DATA_BLOCK "HMI"   // DB2
{ S7_Optimized_Access := 'TRUE' }
VERSION : 0.1
   VAR
      barcode : "Barcode Screen";
      networkHealth : "Network Health Screen";
      partCall : "Part Call Screen";
      screenNumber : Int;
      settings : "Settings";
      simStations : "Simulated Stations";
      tableNav : "Table Nav: HMI";
   END_VAR
BEGIN
END_DATA_BLOCK

DATA_BLOCK "PN Text Library"   // DB3
{ S7_Optimized_Access := 'TRUE' }
VERSION : 0.1
BEGIN
   pnText[0] := WSTRING#'';
   pnText[1] := WSTRING#'11.52.001.0545.000B';
   pnText[2] := WSTRING#'11.52.001.315.000B';
   pnText[3] := WSTRING#'11.52.001.316.001D';
   pnText[4] := WSTRING#'11.54.007.045.015D';
   pnText[5] := WSTRING#'11.54.007.052.007B';
   pnText[6] := WSTRING#'11.54.007.052.008A';
   pnText[7] := WSTRING#'11.54.007.052.009B';
   pnText[8] := WSTRING#'11.54.007.052.010B';
   pnText[9] := WSTRING#'11.54.007.315.026G';
   pnText[10] := WSTRING#'11.54.017.315.001F';
   pnText[11] := WSTRING#'16.08.208.011.010G';
   pnText[12] := WSTRING#'16.08.208.021.020C';
   pnText[13] := WSTRING#'16.08.208.031.020C';
   pnText[14] := WSTRING#'16.08.208.041.000A';
   pnText[15] := WSTRING#'16.08.208.051.000A';
   pnText[16] := WSTRING#'16.08.208.081.010B';
   pnText[17] := WSTRING#'16.08.208.091.000A';
   pnText[18] := WSTRING#'16.08.208.101.010C';
   pnText[19] := WSTRING#'16.08.208.111.000B';
   pnText[20] := WSTRING#'16.08.208.131.010L';
   pnText[21] := WSTRING#'16.08.208.151.010F';
   pnText[22] := WSTRING#'16.08.208.161.020F';
   pnText[23] := WSTRING#'16.08.208.301.000F';
   pnText[24] := WSTRING#'16.08.208.311.000F';
   pnText[25] := WSTRING#'16.08.208.321.000G';
   pnText[26] := WSTRING#'16.08.208.331.000F';
   pnText[27] := WSTRING#'16.08.208.411.030C';
   pnText[28] := WSTRING#'16.08.208.501.000B';
   pnText[29] := WSTRING#'16.08.208.531.020L';
   pnText[30] := WSTRING#'16.08.208.621.010C';
   pnText[31] := WSTRING#'16.08.208.631.000F';
   pnText[32] := WSTRING#'16.08.208.651.010B';
   pnText[33] := WSTRING#'16.08.208.661.000F';
   pnText[34] := WSTRING#'16.08.208.691.010D';
   pnText[35] := WSTRING#'16.08.209.031.010C';
   pnText[36] := WSTRING#'16.08.209.031.030B';
   pnText[37] := WSTRING#'16.08.209.031.050A';
   pnText[38] := WSTRING#'16.08.209.091.010C';
   pnText[39] := WSTRING#'16.08.209.091.030D';
   pnText[40] := WSTRING#'16.08.209.091.060A';
   pnText[41] := WSTRING#'16.08.209.232.010C';
   pnText[42] := WSTRING#'16.08.210.031.010B';
   pnText[43] := WSTRING#'16.08.210.421.010A';
   pnText[44] := WSTRING#'16.08.210.421.020A';
   pnText[45] := WSTRING#'16.08.210.421.030A';
   pnText[46] := WSTRING#'16.08.211.121.000G';
   pnText[47] := WSTRING#'16.08.211.291.000A';
   pnText[48] := WSTRING#'16.08.211.511.020F';
   pnText[49] := WSTRING#'16.08.211.551.000B';
   pnText[50] := WSTRING#'16.08.211.781.000A';
   pnText[51] := WSTRING#'16.08.211.801.010A';
   pnText[52] := WSTRING#'16.08.211.801.020A';
   pnText[53] := WSTRING#'16.08.211.806.020A';
   pnText[54] := WSTRING#'16.08.215.141.010C';
   pnText[55] := WSTRING#'16.08.215.871.010C';
   pnText[56] := WSTRING#'16.08.216.011.030B';
   pnText[57] := WSTRING#'16.08.216.053.000A';
   pnText[58] := WSTRING#'16.08.216.057.001A';
   pnText[59] := WSTRING#'16.08.216.141.010C';
   pnText[60] := WSTRING#'16.08.216.151.010B';
   pnText[61] := WSTRING#'16.08.216.161.020A';
   pnText[62] := WSTRING#'16.08.216.181.010B';
   pnText[63] := WSTRING#'16.08.216.181.090A';
   pnText[64] := WSTRING#'16.08.216.181.100A';
   pnText[65] := WSTRING#'16.08.216.181.110B';
   pnText[66] := WSTRING#'16.08.216.200.050A';
   pnText[67] := WSTRING#'16.08.216.202.080A';
   pnText[68] := WSTRING#'16.08.216.231.000B';
   pnText[69] := WSTRING#'16.08.216.251.000B';
   pnText[70] := WSTRING#'16.08.216.291.000A';
   pnText[71] := WSTRING#'16.08.216.315.000A';
   pnText[72] := WSTRING#'16.08.216.315.001A';
   pnText[73] := WSTRING#'16.08.216.315.002A';
   pnText[74] := WSTRING#'16.08.216.501.000C';
   pnText[75] := WSTRING#'16.08.216.501.010A';
   pnText[76] := WSTRING#'16.08.216.511.000C';
   pnText[77] := WSTRING#'16.08.216.515.008C';
   pnText[78] := WSTRING#'16.08.216.521.000C';
   pnText[79] := WSTRING#'16.08.216.526.002C';
   pnText[80] := WSTRING#'16.08.216.526.009A';
   pnText[81] := WSTRING#'16.08.216.551.000B';
   pnText[82] := WSTRING#'16.08.216.722.001A';
   pnText[83] := WSTRING#'16.08.216.790.001A';
   pnText[84] := WSTRING#'16.08.216.806.020A';
   pnText[85] := WSTRING#'16.08.216.831.020A';
   pnText[86] := WSTRING#'16.08.216.871.010C';
   pnText[87] := WSTRING#'16.08.216.910.020B';
   pnText[88] := WSTRING#'16.08.216.911.000C';
   pnText[89] := WSTRING#'16.08.216.911.000G';
   pnText[90] := WSTRING#'16.08.216.911.000H';
   pnText[91] := WSTRING#'16.08.216.911.030B';
   pnText[92] := WSTRING#'16.08.216.911.040B';
   pnText[93] := WSTRING#'16.08.216.912.050A';
   pnText[94] := WSTRING#'16.08.216.912.060B';
   pnText[95] := WSTRING#'16.08.216.951.010A';
   pnText[96] := WSTRING#'16.08.216.181.020A';
   pnText[97] := WSTRING#'16.08.217.411.080A';
   pnText[98] := WSTRING#'16.08.217.421.010A';
   pnText[99] := WSTRING#'16.08.217.421.130A';
   pnText[100] := WSTRING#'16.18.007.301.010A';
   pnText[101] := WSTRING#'16.18.007.301.020A';
   pnText[102] := WSTRING#'16.18.007.311.010A';
   pnText[103] := WSTRING#'16.18.007.311.020A';
   pnText[104] := WSTRING#'16.18.007.321.010B';
   pnText[105] := WSTRING#'16.18.008.301.010A';
   pnText[106] := WSTRING#'16.18.008.301.020A';
   pnText[107] := WSTRING#'16.18.008.301.030A';
   pnText[108] := WSTRING#'16.18.008.311.010A';
   pnText[109] := WSTRING#'16.18.008.311.020B';
   pnText[110] := WSTRING#'16.18.009.301.010A';
   pnText[111] := WSTRING#'16.18.009.301.020B';
   pnText[112] := WSTRING#'16.18.009.301.030A';
   pnText[113] := WSTRING#'16.18.009.301.040B';
   pnText[114] := WSTRING#'16.18.009.301.050A';
   pnText[115] := WSTRING#'16.18.009.311.010A';
   pnText[116] := WSTRING#'16.18.009.321.010A';
   pnText[117] := WSTRING#'16.18.009.321.020B';
   pnText[118] := WSTRING#'16.18.009.321.030A';
   pnText[119] := WSTRING#'16.18.009.331.030A';
   pnText[120] := WSTRING#'16.18.009.331.050A';
   pnText[121] := WSTRING#'16.18.009.371.010A';
   pnText[122] := WSTRING#'16.18.011.301.010A';
   pnText[123] := WSTRING#'16.18.011.301.020B';
   pnText[124] := WSTRING#'16.18.011.301.030A';
   pnText[125] := WSTRING#'16.18.011.301.040B';
   pnText[126] := WSTRING#'16.18.011.311.020A';
   pnText[127] := WSTRING#'16.18.011.321.010A';
   pnText[128] := WSTRING#'16.18.011.321.020B';
   pnText[129] := WSTRING#'16.18.011.321.030A';
   pnText[130] := WSTRING#'16.18.011.331.010A';
   pnText[131] := WSTRING#'16.18.011.331.020D';
   pnText[132] := WSTRING#'16.18.012.401.010A';
   pnText[133] := WSTRING#'16.18.012.401.020A';
   pnText[134] := WSTRING#'16.18.012.411.010A';
   pnText[135] := WSTRING#'16.18.012.411.020B';
   pnText[136] := WSTRING#'16.18.012.431.010A';
   pnText[137] := WSTRING#'16.18.012.441.010A';
   pnText[138] := WSTRING#'16.18.013.411.010A';
   pnText[139] := WSTRING#'16.18.013.411.020B';
   pnText[140] := WSTRING#'16.18.013.411.030A';
   pnText[141] := WSTRING#'16.18.013.421.010A';
   pnText[142] := WSTRING#'16.18.014.411.010A';
   pnText[143] := WSTRING#'16.18.014.411.030A';
   pnText[144] := WSTRING#'16.18.015.401.010A';
   pnText[145] := WSTRING#'16.18.015.411.010A';
   pnText[146] := WSTRING#'16.18.015.411.020B';
   pnText[147] := WSTRING#'16.18.015.411.030A';
   pnText[148] := WSTRING#'16.18.015.421.010A';
   pnText[149] := WSTRING#'16.18.015.421.020B';
   pnText[150] := WSTRING#'16.18.017.301.010A';
   pnText[151] := WSTRING#'16.18.017.301.020A';
   pnText[152] := WSTRING#'16.18.017.301.030A';
   pnText[153] := WSTRING#'16.18.017.301.040A';
   pnText[154] := WSTRING#'16.18.017.301.050A';
   pnText[155] := WSTRING#'16.18.017.311.010A';
   pnText[156] := WSTRING#'16.18.017.321.010A';
   pnText[157] := WSTRING#'16.18.017.321.020A';
   pnText[158] := WSTRING#'16.18.018.400.000A';
   pnText[159] := WSTRING#'16.18.018.401.010A';
   pnText[160] := WSTRING#'16.18.018.401.020B';
   pnText[161] := WSTRING#'16.18.018.401.030A';
   pnText[162] := WSTRING#'16.18.018.411.010A';
   pnText[163] := WSTRING#'16.18.018.421.010B';
   pnText[164] := WSTRING#'16.32.112.054.041A';
   pnText[165] := WSTRING#'16.32.112.057.010A';
   pnText[166] := WSTRING#'16.32.112.500.060D';
   pnText[167] := WSTRING#'16.32.112.500.090B';
   pnText[168] := WSTRING#'16.32.112.500.100A';
   pnText[169] := WSTRING#'16.32.112.500.120A';
   pnText[170] := WSTRING#'16.32.112.500.150B';
   pnText[171] := WSTRING#'16.32.112.500.160A';
   pnText[172] := WSTRING#'16.32.112.500.220A';
   pnText[173] := WSTRING#'16.32.112.500.300E';
   pnText[174] := WSTRING#'16.32.112.500.520B';
   pnText[175] := WSTRING#'16.32.112.502.050B';
   pnText[176] := WSTRING#'16.32.112.502.060B';
   pnText[177] := WSTRING#'16.32.112.502.070E';
   pnText[178] := WSTRING#'16.32.112.503.210A';
   pnText[179] := WSTRING#'16.32.112.503.220A';
   pnText[180] := WSTRING#'16.32.112.504.060A';
   pnText[181] := WSTRING#'16.32.112.504.070G';
   pnText[182] := WSTRING#'16.32.112.509.050E';
   pnText[183] := WSTRING#'16.32.112.509.070A';
   pnText[184] := WSTRING#'16.32.112.509.080F';
   pnText[185] := WSTRING#'16.32.112.516.110E';
   pnText[186] := WSTRING#'16.32.112.520.300E';
   pnText[187] := WSTRING#'16.32.112.521.010B';
   pnText[188] := WSTRING#'16.32.112.521.020B';
   pnText[189] := WSTRING#'16.32.112.521.030A';
   pnText[190] := WSTRING#'16.32.112.522.040D';
   pnText[191] := WSTRING#'16.32.112.522.050A';
   pnText[192] := WSTRING#'16.32.112.522.130A';
   pnText[193] := WSTRING#'16.32.112.529.010A';
   pnText[194] := WSTRING#'16.32.112.529.020B';
   pnText[195] := WSTRING#'16.32.112.529.030A';
   pnText[196] := WSTRING#'16.32.112.529.050D';
   pnText[197] := WSTRING#'16.32.112.536.010A';
   pnText[198] := WSTRING#'16.32.112.543.020A';
   pnText[199] := WSTRING#'16.32.112.543.210E';
   pnText[200] := WSTRING#'16.32.112.553.010A';
   pnText[201] := WSTRING#'16.32.112.553.020A';
   pnText[202] := WSTRING#'16.32.112.553.100D';
   pnText[203] := WSTRING#'16.32.112.553.220A';
   pnText[204] := WSTRING#'16.32.112.580.020A';
   pnText[205] := WSTRING#'16.32.112.601.030A';
   pnText[206] := WSTRING#'16.32.112.601.040A';
   pnText[207] := WSTRING#'16.32.112.621.010A';
   pnText[208] := WSTRING#'16.32.112.621.020A';
   pnText[209] := WSTRING#'16.32.112.704.000C';
   pnText[210] := WSTRING#'16.32.112.751.000D';
   pnText[211] := WSTRING#'16.32.112.751.001C';
   pnText[212] := WSTRING#'16.32.112.757.000A';
   pnText[213] := WSTRING#'16.32.112.757.001A';
   pnText[214] := WSTRING#'16.32.112.851.000A';
   pnText[215] := WSTRING#'16.32.112.851.001A';
   pnText[216] := WSTRING#'16.32.112.870.000C';
   pnText[217] := WSTRING#'16.32.307.211.150B';
   pnText[218] := WSTRING#'16.32.307.211.170B';
   pnText[219] := WSTRING#'16.32.307.212.320C';
   pnText[220] := WSTRING#'16.32.307.232.300B';
   pnText[221] := WSTRING#'16.32.307.262.300B';
   pnText[222] := WSTRING#'16.32.307.312.310A';
   pnText[223] := WSTRING#'16.32.307.461.160A';
   pnText[224] := WSTRING#'16.32.407.241.150B';
   pnText[225] := WSTRING#'16.32.407.241.170B';
   pnText[226] := WSTRING#'16.32.407.441.160A';
   pnText[227] := WSTRING#'16.32.606.311.010C';
   pnText[228] := WSTRING#'16.32.606.311.040B';
   pnText[229] := WSTRING#'16.32.606.311.050B';
   pnText[230] := WSTRING#'16.32.606.311.060A';
   pnText[231] := WSTRING#'16.32.606.311.070A';
   pnText[232] := WSTRING#'16.32.606.321.010B';
   pnText[233] := WSTRING#'16.32.606.321.030B';
   pnText[234] := WSTRING#'16.32.706.311.010C';
   pnText[235] := WSTRING#'16.32.706.311.020B';
   pnText[236] := WSTRING#'16.32.706.311.040B';
   pnText[237] := WSTRING#'16.32.706.311.050B';
   pnText[238] := WSTRING#'16.32.706.321.010B';
   pnText[239] := WSTRING#'16.32.706.321.030B';
   pnText[240] := WSTRING#'16.32.706.401.040A';
   pnText[241] := WSTRING#'16.32.706.401.050A';
   pnText[242] := WSTRING#'16.32.806.502.080A';
   pnText[243] := WSTRING#'DUNNAGE';
   pnText[244] := WSTRING#'PEANUTS';
   pnText[245] := WSTRING#'RINGS CART';
END_DATA_BLOCK

DATA_BLOCK "LED Sign"   // DB4
{ S7_Optimized_Access := 'TRUE' }
VERSION : 0.1
   VAR
      request : "LED Sign Data";
   END_VAR
BEGIN
END_DATA_BLOCK

DATA_BLOCK "Recipe Buffer"   // DB5
{ S7_Optimized_Access := 'TRUE' }
VERSION : 0.1
BEGIN
END_DATA_BLOCK

DATA_BLOCK "HMI Stations"   // DB6
{ S7_Optimized_Access := 'TRUE' }
VERSION : 0.1
   VAR
      me : Array[0.."hmiStnCount"] of "HMIS: Compressed";
   END_VAR
BEGIN
END_DATA_BLOCK

DATA_BLOCK "Stations"   // DB10
{ S7_Optimized_Access := 'TRUE' }
VERSION : 0.1
BEGIN
   stn[0].id.dropZone := 1;
   stn[0].id.lineName := WSTRING#'VOLVO 16';
   stn[0].ioData.kp8.output := 16#0000_0000;
   stn[0].ioData.stkLight := 16#0000_0000;
   stn[0].wipData."name" := WSTRING#'';
   stn[1].id.dropZone := 2;
   stn[1].id.lineName := WSTRING#'VOLVO 16';
   stn[1].ioData.kp8.output := 16#0000_0000;
   stn[1].ioData.stkLight := 16#0000_0000;
   stn[1].wipData."name" := WSTRING#'';
   stn[2].id.dropZone := 3;
   stn[2].id.lineName := WSTRING#'VOLVO 16';
   stn[2].ioData.kp8.output := 16#0000_0000;
   stn[2].ioData.stkLight := 16#0000_0000;
   stn[2].wipData."name" := WSTRING#'';
   stn[3].id.dropZone := 4;
   stn[3].id.lineName := WSTRING#'VOLVO 16';
   stn[3].ioData.kp8.output := 16#0000_0000;
   stn[3].ioData.stkLight := 16#0000_0000;
   stn[3].wipData."name" := WSTRING#'';
   stn[4].id.lineName := WSTRING#'';
   stn[4].ioData.kp8.output := 16#0000_0000;
   stn[4].ioData.stkLight := 16#0000_0000;
   stn[4].wipData."name" := WSTRING#'';
   stn[5].id.lineName := WSTRING#'';
   stn[5].ioData.kp8.output := 16#0000_0000;
   stn[5].ioData.stkLight := 16#0000_0000;
   stn[5].wipData."name" := WSTRING#'';
   stn[6].id.lineName := WSTRING#'';
   stn[6].ioData.kp8.output := 16#0000_0000;
   stn[6].ioData.stkLight := 16#0000_0000;
   stn[6].wipData."name" := WSTRING#'';
   stn[7].id.lineName := WSTRING#'';
   stn[7].ioData.kp8.output := 16#0000_0000;
   stn[7].ioData.stkLight := 16#0000_0000;
   stn[7].wipData."name" := WSTRING#'';
   stn[8].id.lineName := WSTRING#'';
   stn[8].ioData.kp8.output := 16#0000_0000;
   stn[8].ioData.stkLight := 16#0000_0000;
   stn[8].wipData."name" := WSTRING#'';
   stn[9].id.lineName := WSTRING#'';
   stn[9].ioData.kp8.output := 16#0000_0000;
   stn[9].ioData.stkLight := 16#0000_0000;
   stn[9].wipData."name" := WSTRING#'';
   stn[10].id.lineName := WSTRING#'';
   stn[10].ioData.kp8.output := 16#0000_0000;
   stn[10].ioData.stkLight := 16#0000_0000;
   stn[10].wipData."name" := WSTRING#'';
   stn[11].id.lineName := WSTRING#'';
   stn[11].ioData.kp8.output := 16#0000_0000;
   stn[11].ioData.stkLight := 16#0000_0000;
   stn[11].wipData."name" := WSTRING#'';
   stn[12].id.lineName := WSTRING#'';
   stn[12].ioData.kp8.output := 16#0000_0000;
   stn[12].ioData.stkLight := 16#0000_0000;
   stn[12].wipData."name" := WSTRING#'';
   stn[13].id.lineName := WSTRING#'';
   stn[13].ioData.kp8.output := 16#0000_0000;
   stn[13].ioData.stkLight := 16#0000_0000;
   stn[13].wipData."name" := WSTRING#'';
   stn[14].id.lineName := WSTRING#'';
   stn[14].ioData.kp8.output := 16#0000_0000;
   stn[14].ioData.stkLight := 16#0000_0000;
   stn[14].wipData."name" := WSTRING#'';
   stn[15].id.lineName := WSTRING#'';
   stn[15].ioData.kp8.output := 16#0000_0000;
   stn[15].ioData.stkLight := 16#0000_0000;
   stn[15].wipData."name" := WSTRING#'';
   stn[16].id.lineName := WSTRING#'';
   stn[16].ioData.kp8.output := 16#0000_0000;
   stn[16].ioData.stkLight := 16#0000_0000;
   stn[16].wipData."name" := WSTRING#'';
   stn[17].id.lineName := WSTRING#'';
   stn[17].ioData.kp8.output := 16#0000_0000;
   stn[17].ioData.stkLight := 16#0000_0000;
   stn[17].wipData."name" := WSTRING#'';
   stn[18].id.lineName := WSTRING#'';
   stn[18].ioData.kp8.output := 16#0000_0000;
   stn[18].ioData.stkLight := 16#0000_0000;
   stn[18].wipData."name" := WSTRING#'';
   stn[19].id.lineName := WSTRING#'';
   stn[19].ioData.kp8.output := 16#0000_0000;
   stn[19].ioData.stkLight := 16#0000_0000;
   stn[19].wipData."name" := WSTRING#'';
   stn[20].id.lineName := WSTRING#'';
   stn[20].ioData.kp8.output := 16#0000_0000;
   stn[20].ioData.stkLight := 16#0000_0000;
   stn[20].wipData."name" := WSTRING#'';
   stn[21].id.lineName := WSTRING#'';
   stn[21].ioData.kp8.output := 16#0000_0000;
   stn[21].ioData.stkLight := 16#0000_0000;
   stn[21].wipData."name" := WSTRING#'';
   stn[22].id.lineName := WSTRING#'';
   stn[22].ioData.kp8.output := 16#0000_0000;
   stn[22].ioData.stkLight := 16#0000_0000;
   stn[22].wipData."name" := WSTRING#'';
   stn[23].id.lineName := WSTRING#'';
   stn[23].ioData.kp8.output := 16#0000_0000;
   stn[23].ioData.stkLight := 16#0000_0000;
   stn[23].wipData."name" := WSTRING#'';
   stn[24].id.lineName := WSTRING#'';
   stn[24].ioData.kp8.output := 16#0000_0000;
   stn[24].ioData.stkLight := 16#0000_0000;
   stn[24].wipData."name" := WSTRING#'';
   stn[25].id.lineName := WSTRING#'';
   stn[25].ioData.kp8.output := 16#0000_0000;
   stn[25].ioData.stkLight := 16#0000_0000;
   stn[25].wipData."name" := WSTRING#'';
   stn[26].id.lineName := WSTRING#'';
   stn[26].ioData.kp8.output := 16#0000_0000;
   stn[26].ioData.stkLight := 16#0000_0000;
   stn[26].wipData."name" := WSTRING#'';
   stn[27].id.lineName := WSTRING#'';
   stn[27].ioData.kp8.output := 16#0000_0000;
   stn[27].ioData.stkLight := 16#0000_0000;
   stn[27].wipData."name" := WSTRING#'';
   stn[28].id.lineName := WSTRING#'';
   stn[28].ioData.kp8.output := 16#0000_0000;
   stn[28].ioData.stkLight := 16#0000_0000;
   stn[28].wipData."name" := WSTRING#'';
   stn[29].id.lineName := WSTRING#'';
   stn[29].ioData.kp8.output := 16#0000_0000;
   stn[29].ioData.stkLight := 16#0000_0000;
   stn[29].wipData."name" := WSTRING#'';
   stn[30].id.lineName := WSTRING#'';
   stn[30].ioData.kp8.output := 16#0000_0000;
   stn[30].ioData.stkLight := 16#0000_0000;
   stn[30].wipData."name" := WSTRING#'';
   stn[31].id.lineName := WSTRING#'';
   stn[31].ioData.kp8.output := 16#0000_0000;
   stn[31].ioData.stkLight := 16#0000_0000;
   stn[31].wipData."name" := WSTRING#'';
   stn[32].id.lineName := WSTRING#'';
   stn[32].ioData.kp8.output := 16#0000_0000;
   stn[32].ioData.stkLight := 16#0000_0000;
   stn[32].wipData."name" := WSTRING#'';
   stn[33].id.lineName := WSTRING#'';
   stn[33].ioData.kp8.output := 16#0000_0000;
   stn[33].ioData.stkLight := 16#0000_0000;
   stn[33].wipData."name" := WSTRING#'';
   stn[34].id.lineName := WSTRING#'';
   stn[34].ioData.kp8.output := 16#0000_0000;
   stn[34].ioData.stkLight := 16#0000_0000;
   stn[34].wipData."name" := WSTRING#'';
   stn[35].id.lineName := WSTRING#'';
   stn[35].ioData.kp8.output := 16#0000_0000;
   stn[35].ioData.stkLight := 16#0000_0000;
   stn[35].wipData."name" := WSTRING#'';
   stn[36].id.lineName := WSTRING#'';
   stn[36].ioData.kp8.output := 16#0000_0000;
   stn[36].ioData.stkLight := 16#0000_0000;
   stn[36].wipData."name" := WSTRING#'';
   stn[37].id.lineName := WSTRING#'';
   stn[37].ioData.kp8.output := 16#0000_0000;
   stn[37].ioData.stkLight := 16#0000_0000;
   stn[37].wipData."name" := WSTRING#'';
   stn[38].id.lineName := WSTRING#'';
   stn[38].ioData.kp8.output := 16#0000_0000;
   stn[38].ioData.stkLight := 16#0000_0000;
   stn[38].wipData."name" := WSTRING#'';
END_DATA_BLOCK

DATA_BLOCK "Part Requests"   // DB11
{ S7_Optimized_Access := 'TRUE' }
VERSION : 0.1
BEGIN
END_DATA_BLOCK

DATA_BLOCK "PN Code Library"   // DB12
{ S7_Optimized_Access := 'TRUE' }
VERSION : 0.1
BEGIN
   stn[0].wipBtn[0,0] := 0;
   stn[0].wipBtn[0,1] := 0;
   stn[0].wipBtn[0,2] := 0;
   stn[0].wipBtn[0,4] := 0;
   stn[0].wipBtn[0,5] := 0;
   stn[0].wipBtn[0,6] := 0;
   stn[0].wipBtn[1,0] := 0;
   stn[0].wipBtn[1,1] := 0;
   stn[0].wipBtn[1,2] := 0;
   stn[0].wipBtn[1,3] := 0;
   stn[0].wipBtn[1,4] := 0;
   stn[0].wipBtn[1,5] := 0;
   stn[0].wipBtn[1,6] := 0;
   stn[0].wipBtn[1,7] := 0;
   stn[0].wipBtn[2,0] := 0;
   stn[0].wipBtn[2,1] := 0;
   stn[0].wipBtn[2,2] := 0;
   stn[0].wipBtn[2,3] := 0;
   stn[0].wipBtn[2,4] := 0;
   stn[0].wipBtn[2,5] := 0;
   stn[0].wipBtn[2,6] := 0;
   stn[0].wipBtn[2,7] := 0;
   stn[0].wipBtn[3,0] := 0;
   stn[0].wipBtn[3,1] := 0;
   stn[0].wipBtn[3,2] := 0;
   stn[0].wipBtn[3,3] := 0;
   stn[0].wipBtn[3,4] := 0;
   stn[0].wipBtn[3,5] := 0;
   stn[0].wipBtn[3,6] := 0;
   stn[0].wipBtn[3,7] := 0;
   stn[0].wipBtn[4,0] := 0;
   stn[0].wipBtn[4,1] := 0;
   stn[0].wipBtn[4,2] := 0;
   stn[0].wipBtn[4,3] := 0;
   stn[0].wipBtn[4,4] := 0;
   stn[0].wipBtn[4,5] := 0;
   stn[0].wipBtn[4,6] := 0;
   stn[0].wipBtn[4,7] := 0;
   stn[0].wipBtn[5,0] := 0;
   stn[0].wipBtn[5,1] := 0;
   stn[0].wipBtn[5,2] := 0;
   stn[0].wipBtn[5,3] := 0;
   stn[0].wipBtn[5,4] := 0;
   stn[0].wipBtn[5,5] := 0;
   stn[0].wipBtn[5,6] := 0;
   stn[0].wipBtn[5,7] := 0;
   stn[0].wipBtn[6,0] := 0;
   stn[0].wipBtn[6,1] := 0;
   stn[0].wipBtn[6,2] := 0;
   stn[0].wipBtn[6,3] := 0;
   stn[0].wipBtn[6,4] := 0;
   stn[0].wipBtn[6,5] := 0;
   stn[0].wipBtn[6,6] := 0;
   stn[0].wipBtn[6,7] := 0;
   stn[0].wipBtn[7,0] := 0;
   stn[0].wipBtn[7,1] := 0;
   stn[0].wipBtn[7,2] := 0;
   stn[0].wipBtn[7,3] := 0;
   stn[0].wipBtn[7,4] := 0;
   stn[0].wipBtn[7,5] := 0;
   stn[0].wipBtn[7,6] := 0;
   stn[0].wipBtn[7,7] := 0;
   stn[0].wipBtn[8,0] := 0;
   stn[0].wipBtn[8,1] := 0;
   stn[0].wipBtn[8,2] := 0;
   stn[0].wipBtn[8,3] := 0;
   stn[0].wipBtn[8,4] := 0;
   stn[0].wipBtn[8,5] := 0;
   stn[0].wipBtn[8,6] := 0;
   stn[0].wipBtn[8,7] := 0;
   stn[0].wipBtn[9,0] := 0;
   stn[0].wipBtn[9,1] := 0;
   stn[0].wipBtn[9,2] := 0;
   stn[0].wipBtn[9,3] := 0;
   stn[0].wipBtn[9,4] := 0;
   stn[0].wipBtn[9,5] := 0;
   stn[0].wipBtn[9,6] := 0;
   stn[0].wipBtn[9,7] := 0;
   stn[0].wipBtn[10,0] := 0;
   stn[0].wipBtn[10,1] := 0;
   stn[0].wipBtn[10,2] := 0;
   stn[0].wipBtn[10,3] := 0;
   stn[0].wipBtn[10,4] := 0;
   stn[0].wipBtn[10,5] := 0;
   stn[0].wipBtn[10,6] := 0;
   stn[0].wipBtn[10,7] := 0;
   stn[0].wipBtn[11,0] := 0;
   stn[0].wipBtn[11,1] := 0;
   stn[0].wipBtn[11,2] := 0;
   stn[0].wipBtn[11,3] := 0;
   stn[0].wipBtn[11,4] := 0;
   stn[0].wipBtn[11,5] := 0;
   stn[0].wipBtn[11,6] := 0;
   stn[0].wipBtn[11,7] := 0;
   stn[0].wipBtn[12,0] := 0;
   stn[0].wipBtn[12,1] := 0;
   stn[0].wipBtn[12,2] := 0;
   stn[0].wipBtn[12,3] := 0;
   stn[0].wipBtn[12,4] := 0;
   stn[0].wipBtn[12,5] := 0;
   stn[0].wipBtn[12,6] := 0;
   stn[0].wipBtn[12,7] := 0;
   stn[0].wipBtn[13,0] := 0;
   stn[0].wipBtn[13,1] := 0;
   stn[0].wipBtn[13,2] := 0;
   stn[0].wipBtn[13,3] := 0;
   stn[0].wipBtn[13,4] := 0;
   stn[0].wipBtn[13,5] := 0;
   stn[0].wipBtn[13,6] := 0;
   stn[0].wipBtn[13,7] := 0;
   stn[0].wipBtn[14,0] := 0;
   stn[0].wipBtn[14,1] := 0;
   stn[0].wipBtn[14,2] := 0;
   stn[0].wipBtn[14,3] := 0;
   stn[0].wipBtn[14,4] := 0;
   stn[0].wipBtn[14,5] := 0;
   stn[0].wipBtn[14,6] := 0;
   stn[0].wipBtn[14,7] := 0;
   stn[0].wipBtn[15,0] := 0;
   stn[0].wipBtn[15,1] := 0;
   stn[0].wipBtn[15,2] := 0;
   stn[0].wipBtn[15,3] := 0;
   stn[0].wipBtn[15,4] := 0;
   stn[0].wipBtn[15,5] := 0;
   stn[0].wipBtn[15,6] := 0;
   stn[0].wipBtn[15,7] := 0;
   stn[0].wipBtn[16,0] := 0;
   stn[0].wipBtn[16,1] := 0;
   stn[0].wipBtn[16,2] := 0;
   stn[0].wipBtn[16,3] := 0;
   stn[0].wipBtn[16,4] := 0;
   stn[0].wipBtn[16,5] := 0;
   stn[0].wipBtn[16,6] := 0;
   stn[0].wipBtn[16,7] := 0;
   stn[0].wipBtn[17,0] := 0;
   stn[0].wipBtn[17,1] := 0;
   stn[0].wipBtn[17,2] := 0;
   stn[0].wipBtn[17,3] := 0;
   stn[0].wipBtn[17,4] := 0;
   stn[0].wipBtn[17,5] := 0;
   stn[0].wipBtn[17,6] := 0;
   stn[0].wipBtn[17,7] := 0;
   stn[0].wipBtn[18,0] := 0;
   stn[0].wipBtn[18,1] := 0;
   stn[0].wipBtn[18,2] := 0;
   stn[0].wipBtn[18,3] := 0;
   stn[0].wipBtn[18,4] := 0;
   stn[0].wipBtn[18,5] := 0;
   stn[0].wipBtn[18,6] := 0;
   stn[0].wipBtn[18,7] := 0;
   stn[0].wipBtn[19,0] := 0;
   stn[0].wipBtn[19,1] := 0;
   stn[0].wipBtn[19,2] := 0;
   stn[0].wipBtn[19,3] := 0;
   stn[0].wipBtn[19,4] := 0;
   stn[0].wipBtn[19,5] := 0;
   stn[0].wipBtn[19,6] := 0;
   stn[0].wipBtn[19,7] := 0;
   stn[0].wipBtn[20,0] := 0;
   stn[0].wipBtn[20,1] := 0;
   stn[0].wipBtn[20,2] := 0;
   stn[0].wipBtn[20,3] := 0;
   stn[0].wipBtn[20,4] := 0;
   stn[0].wipBtn[20,5] := 0;
   stn[0].wipBtn[20,6] := 0;
   stn[0].wipBtn[20,7] := 0;
   stn[0].wipBtn[21,0] := 0;
   stn[0].wipBtn[21,1] := 0;
   stn[0].wipBtn[21,2] := 0;
   stn[0].wipBtn[21,3] := 0;
   stn[0].wipBtn[21,4] := 0;
   stn[0].wipBtn[21,5] := 0;
   stn[0].wipBtn[21,6] := 0;
   stn[0].wipBtn[21,7] := 0;
   stn[0].wipBtn[22,0] := 0;
   stn[0].wipBtn[22,1] := 0;
   stn[0].wipBtn[22,2] := 0;
   stn[0].wipBtn[22,3] := 0;
   stn[0].wipBtn[22,4] := 0;
   stn[0].wipBtn[22,5] := 0;
   stn[0].wipBtn[22,6] := 0;
   stn[0].wipBtn[22,7] := 0;
   stn[0].wipBtn[23,0] := 0;
   stn[0].wipBtn[23,1] := 0;
   stn[0].wipBtn[23,2] := 0;
   stn[0].wipBtn[23,3] := 0;
   stn[0].wipBtn[23,4] := 0;
   stn[0].wipBtn[23,5] := 0;
   stn[0].wipBtn[23,6] := 0;
   stn[0].wipBtn[23,7] := 0;
   stn[0].wipBtn[24,0] := 0;
   stn[0].wipBtn[24,1] := 0;
   stn[0].wipBtn[24,2] := 0;
   stn[0].wipBtn[24,3] := 0;
   stn[0].wipBtn[24,4] := 0;
   stn[0].wipBtn[24,5] := 0;
   stn[0].wipBtn[24,6] := 0;
   stn[0].wipBtn[24,7] := 0;
   stn[0].wipBtn[25,0] := 0;
   stn[0].wipBtn[25,1] := 0;
   stn[0].wipBtn[25,2] := 0;
   stn[0].wipBtn[25,3] := 0;
   stn[0].wipBtn[25,4] := 0;
   stn[0].wipBtn[25,5] := 0;
   stn[0].wipBtn[25,6] := 0;
   stn[0].wipBtn[25,7] := 0;
   stn[0].wipBtn[26,0] := 0;
   stn[0].wipBtn[26,1] := 0;
   stn[0].wipBtn[26,2] := 0;
   stn[0].wipBtn[26,3] := 0;
   stn[0].wipBtn[26,4] := 0;
   stn[0].wipBtn[26,5] := 0;
   stn[0].wipBtn[26,6] := 0;
   stn[0].wipBtn[26,7] := 0;
   stn[0].wipBtn[27,0] := 0;
   stn[0].wipBtn[27,1] := 0;
   stn[0].wipBtn[27,2] := 0;
   stn[0].wipBtn[27,3] := 0;
   stn[0].wipBtn[27,4] := 0;
   stn[0].wipBtn[27,5] := 0;
   stn[0].wipBtn[27,6] := 0;
   stn[0].wipBtn[27,7] := 0;
   stn[0].wipBtn[28,0] := 0;
   stn[0].wipBtn[28,1] := 0;
   stn[0].wipBtn[28,2] := 0;
   stn[0].wipBtn[28,3] := 0;
   stn[0].wipBtn[28,4] := 0;
   stn[0].wipBtn[28,5] := 0;
   stn[0].wipBtn[28,6] := 0;
   stn[0].wipBtn[28,7] := 0;
   stn[0].wipBtn[29,0] := 0;
   stn[0].wipBtn[29,1] := 0;
   stn[0].wipBtn[29,2] := 0;
   stn[0].wipBtn[29,3] := 0;
   stn[0].wipBtn[29,4] := 0;
   stn[0].wipBtn[29,5] := 0;
   stn[0].wipBtn[29,6] := 0;
   stn[0].wipBtn[29,7] := 0;
   stn[0].wipBtn[30,0] := 0;
   stn[0].wipBtn[30,1] := 0;
   stn[0].wipBtn[30,2] := 0;
   stn[0].wipBtn[30,3] := 0;
   stn[0].wipBtn[30,4] := 0;
   stn[0].wipBtn[30,5] := 0;
   stn[0].wipBtn[30,6] := 0;
   stn[0].wipBtn[30,7] := 0;
   stn[0].wipBtn[31,0] := 0;
   stn[0].wipBtn[31,1] := 0;
   stn[0].wipBtn[31,2] := 0;
   stn[0].wipBtn[31,3] := 0;
   stn[0].wipBtn[31,4] := 0;
   stn[0].wipBtn[31,5] := 0;
   stn[0].wipBtn[31,6] := 0;
   stn[0].wipBtn[31,7] := 0;
   stn[0].wipBtn[32,0] := 0;
   stn[0].wipBtn[32,1] := 0;
   stn[0].wipBtn[32,2] := 0;
   stn[0].wipBtn[32,3] := 0;
   stn[0].wipBtn[32,4] := 0;
   stn[0].wipBtn[32,5] := 0;
   stn[0].wipBtn[32,6] := 0;
   stn[0].wipBtn[32,7] := 0;
   stn[0].wipBtn[33,0] := 0;
   stn[0].wipBtn[33,1] := 0;
   stn[0].wipBtn[33,2] := 0;
   stn[0].wipBtn[33,3] := 0;
   stn[0].wipBtn[33,4] := 0;
   stn[0].wipBtn[33,5] := 0;
   stn[0].wipBtn[33,6] := 0;
   stn[0].wipBtn[33,7] := 0;
   stn[0].wipBtn[34,0] := 0;
   stn[0].wipBtn[34,1] := 0;
   stn[0].wipBtn[34,2] := 0;
   stn[0].wipBtn[34,3] := 0;
   stn[0].wipBtn[34,4] := 0;
   stn[0].wipBtn[34,5] := 0;
   stn[0].wipBtn[34,6] := 0;
   stn[0].wipBtn[34,7] := 0;
   stn[0].wipBtn[35,0] := 0;
   stn[0].wipBtn[35,1] := 0;
   stn[0].wipBtn[35,2] := 0;
   stn[0].wipBtn[35,3] := 0;
   stn[0].wipBtn[35,4] := 0;
   stn[0].wipBtn[35,5] := 0;
   stn[0].wipBtn[35,6] := 0;
   stn[0].wipBtn[35,7] := 0;
   stn[0].wipBtn[36,0] := 0;
   stn[0].wipBtn[36,1] := 0;
   stn[0].wipBtn[36,2] := 0;
   stn[0].wipBtn[36,3] := 0;
   stn[0].wipBtn[36,4] := 0;
   stn[0].wipBtn[36,5] := 0;
   stn[0].wipBtn[36,6] := 0;
   stn[0].wipBtn[36,7] := 0;
   stn[0].wipBtn[37,0] := 0;
   stn[0].wipBtn[37,1] := 0;
   stn[0].wipBtn[37,2] := 0;
   stn[0].wipBtn[37,3] := 0;
   stn[0].wipBtn[37,4] := 0;
   stn[0].wipBtn[37,5] := 0;
   stn[0].wipBtn[37,6] := 0;
   stn[0].wipBtn[37,7] := 0;
   stn[0].wipBtn[38,0] := 0;
   stn[0].wipBtn[38,1] := 0;
   stn[0].wipBtn[38,2] := 0;
   stn[0].wipBtn[38,3] := 0;
   stn[0].wipBtn[38,4] := 0;
   stn[0].wipBtn[38,5] := 0;
   stn[0].wipBtn[38,6] := 0;
   stn[0].wipBtn[38,7] := 0;
   stn[0].wipBtn[39,0] := 0;
   stn[0].wipBtn[39,1] := 0;
   stn[0].wipBtn[39,2] := 0;
   stn[0].wipBtn[39,3] := 0;
   stn[0].wipBtn[39,4] := 0;
   stn[0].wipBtn[39,5] := 0;
   stn[0].wipBtn[39,6] := 0;
   stn[0].wipBtn[39,7] := 0;
   stn[0].wipBtn[40,0] := 0;
   stn[0].wipBtn[40,1] := 0;
   stn[0].wipBtn[40,2] := 0;
   stn[0].wipBtn[40,3] := 0;
   stn[0].wipBtn[40,4] := 0;
   stn[0].wipBtn[40,5] := 0;
   stn[0].wipBtn[40,6] := 0;
   stn[0].wipBtn[40,7] := 0;
   stn[0].wipBtn[41,0] := 0;
   stn[0].wipBtn[41,1] := 0;
   stn[0].wipBtn[41,2] := 0;
   stn[0].wipBtn[41,3] := 0;
   stn[0].wipBtn[41,4] := 0;
   stn[0].wipBtn[41,5] := 0;
   stn[0].wipBtn[41,6] := 0;
   stn[0].wipBtn[41,7] := 0;
   stn[0].wipBtn[42,0] := 0;
   stn[0].wipBtn[42,1] := 0;
   stn[0].wipBtn[42,2] := 0;
   stn[0].wipBtn[42,3] := 0;
   stn[0].wipBtn[42,4] := 0;
   stn[0].wipBtn[42,5] := 0;
   stn[0].wipBtn[42,6] := 0;
   stn[0].wipBtn[42,7] := 0;
   stn[0].wipBtn[43,0] := 0;
   stn[0].wipBtn[43,1] := 0;
   stn[0].wipBtn[43,2] := 0;
   stn[0].wipBtn[43,3] := 0;
   stn[0].wipBtn[43,4] := 0;
   stn[0].wipBtn[43,5] := 0;
   stn[0].wipBtn[43,6] := 0;
   stn[0].wipBtn[43,7] := 0;
   stn[0].wipBtn[44,0] := 0;
   stn[0].wipBtn[44,1] := 0;
   stn[0].wipBtn[44,2] := 0;
   stn[0].wipBtn[44,3] := 0;
   stn[0].wipBtn[44,4] := 0;
   stn[0].wipBtn[44,5] := 0;
   stn[0].wipBtn[44,6] := 0;
   stn[0].wipBtn[44,7] := 0;
   stn[0].wipBtn[45,0] := 0;
   stn[0].wipBtn[45,1] := 0;
   stn[0].wipBtn[45,2] := 0;
   stn[0].wipBtn[45,3] := 0;
   stn[0].wipBtn[45,4] := 0;
   stn[0].wipBtn[45,5] := 0;
   stn[0].wipBtn[45,6] := 0;
   stn[0].wipBtn[45,7] := 0;
   stn[0].wipBtn[46,0] := 0;
   stn[0].wipBtn[46,1] := 0;
   stn[0].wipBtn[46,2] := 0;
   stn[0].wipBtn[46,3] := 0;
   stn[0].wipBtn[46,4] := 0;
   stn[0].wipBtn[46,5] := 0;
   stn[0].wipBtn[46,6] := 0;
   stn[0].wipBtn[46,7] := 0;
   stn[0].wipBtn[47,0] := 0;
   stn[0].wipBtn[47,1] := 0;
   stn[0].wipBtn[47,2] := 0;
   stn[0].wipBtn[47,3] := 0;
   stn[0].wipBtn[47,4] := 0;
   stn[0].wipBtn[47,5] := 0;
   stn[0].wipBtn[47,6] := 0;
   stn[0].wipBtn[47,7] := 0;
   stn[0].wipBtn[48,0] := 0;
   stn[0].wipBtn[48,1] := 0;
   stn[0].wipBtn[48,2] := 0;
   stn[0].wipBtn[48,3] := 0;
   stn[0].wipBtn[48,4] := 0;
   stn[0].wipBtn[48,5] := 0;
   stn[0].wipBtn[48,6] := 0;
   stn[0].wipBtn[48,7] := 0;
   stn[0].wipBtn[49,0] := 0;
   stn[0].wipBtn[49,1] := 0;
   stn[0].wipBtn[49,2] := 0;
   stn[0].wipBtn[49,3] := 0;
   stn[0].wipBtn[49,4] := 0;
   stn[0].wipBtn[49,5] := 0;
   stn[0].wipBtn[49,6] := 0;
   stn[0].wipBtn[49,7] := 0;
   stn[1].wipBtn[0,0] := 0;
   stn[1].wipBtn[0,1] := 0;
   stn[1].wipBtn[0,3] := 200000;
   stn[1].wipBtn[0,4] := 0;
   stn[1].wipBtn[0,5] := 0;
   stn[1].wipBtn[0,6] := 180000;
   stn[1].wipBtn[1,0] := 0;
   stn[1].wipBtn[1,1] := 0;
   stn[1].wipBtn[1,2] := 0;
   stn[1].wipBtn[1,3] := 0;
   stn[1].wipBtn[1,4] := 0;
   stn[1].wipBtn[1,5] := 0;
   stn[1].wipBtn[1,6] := 0;
   stn[1].wipBtn[1,7] := 0;
   stn[1].wipBtn[2,0] := 0;
   stn[1].wipBtn[2,1] := 0;
   stn[1].wipBtn[2,2] := 0;
   stn[1].wipBtn[2,3] := 0;
   stn[1].wipBtn[2,4] := 0;
   stn[1].wipBtn[2,5] := 0;
   stn[1].wipBtn[2,6] := 0;
   stn[1].wipBtn[2,7] := 0;
   stn[1].wipBtn[3,0] := 0;
   stn[1].wipBtn[3,1] := 0;
   stn[1].wipBtn[3,2] := 0;
   stn[1].wipBtn[3,3] := 0;
   stn[1].wipBtn[3,4] := 0;
   stn[1].wipBtn[3,5] := 0;
   stn[1].wipBtn[3,6] := 0;
   stn[1].wipBtn[3,7] := 0;
   stn[1].wipBtn[4,0] := 0;
   stn[1].wipBtn[4,1] := 0;
   stn[1].wipBtn[4,2] := 0;
   stn[1].wipBtn[4,3] := 0;
   stn[1].wipBtn[4,4] := 0;
   stn[1].wipBtn[4,5] := 0;
   stn[1].wipBtn[4,6] := 0;
   stn[1].wipBtn[4,7] := 0;
   stn[1].wipBtn[5,0] := 0;
   stn[1].wipBtn[5,1] := 0;
   stn[1].wipBtn[5,2] := 0;
   stn[1].wipBtn[5,3] := 0;
   stn[1].wipBtn[5,4] := 0;
   stn[1].wipBtn[5,5] := 0;
   stn[1].wipBtn[5,6] := 0;
   stn[1].wipBtn[5,7] := 0;
   stn[1].wipBtn[6,0] := 0;
   stn[1].wipBtn[6,1] := 0;
   stn[1].wipBtn[6,2] := 0;
   stn[1].wipBtn[6,3] := 0;
   stn[1].wipBtn[6,4] := 0;
   stn[1].wipBtn[6,5] := 0;
   stn[1].wipBtn[6,6] := 0;
   stn[1].wipBtn[6,7] := 0;
   stn[1].wipBtn[7,0] := 0;
   stn[1].wipBtn[7,1] := 0;
   stn[1].wipBtn[7,2] := 0;
   stn[1].wipBtn[7,3] := 0;
   stn[1].wipBtn[7,4] := 0;
   stn[1].wipBtn[7,5] := 0;
   stn[1].wipBtn[7,6] := 0;
   stn[1].wipBtn[7,7] := 0;
   stn[1].wipBtn[8,0] := 0;
   stn[1].wipBtn[8,1] := 0;
   stn[1].wipBtn[8,2] := 0;
   stn[1].wipBtn[8,3] := 0;
   stn[1].wipBtn[8,4] := 0;
   stn[1].wipBtn[8,5] := 0;
   stn[1].wipBtn[8,6] := 0;
   stn[1].wipBtn[8,7] := 0;
   stn[1].wipBtn[9,0] := 0;
   stn[1].wipBtn[9,1] := 0;
   stn[1].wipBtn[9,2] := 0;
   stn[1].wipBtn[9,3] := 0;
   stn[1].wipBtn[9,4] := 0;
   stn[1].wipBtn[9,5] := 0;
   stn[1].wipBtn[9,6] := 0;
   stn[1].wipBtn[9,7] := 0;
   stn[1].wipBtn[10,0] := 0;
   stn[1].wipBtn[10,1] := 0;
   stn[1].wipBtn[10,2] := 0;
   stn[1].wipBtn[10,3] := 0;